REGION Network 6: Programmnummer gültig an den Schäumroboter
   //----
         L     #AB_KUKA_PGNO;
         T     #Prog_Nummer;
   //----
   // Partitätsbit auswerten
   //----
         X     #Temp_IO_Status.Output_To_Robot.A_SPS_PGNO.%X0;
         X     #Temp_IO_Status.Output_To_Robot.A_SPS_PGNO.%X1;
         X     #Temp_IO_Status.Output_To_Robot.A_SPS_PGNO.%X2;
         X     #Temp_IO_Status.Output_To_Robot.A_SPS_PGNO.%X3;
         X     #Temp_IO_Status.Output_To_Robot.A_SPS_PGNO.%X4;
         X     #Temp_IO_Status.Output_To_Robot.A_SPS_PGNO.%X5;
         X     #Temp_IO_Status.Output_To_Robot.A_SPS_PGNO.%X6;
         X     #Temp_IO_Status.Output_To_Robot.A_SPS_PGNO.%X7;
         =     #Temp_IO_Status.Output_To_Robot.A_SPS_PARITY;
   //----
   // Programmnummer an KUKA ablöschen, sobald sie erkannt wurde
   //----
         O(;
         A     #Temp_IO_Status.Input_From_Robot.E_KRC_PGNO_REQ;
         FN    #Temp_IO_Status.FHM_PRG_laeuft;
         );
         ON    #Temp_IO_Status.Input_From_Robot.E_KRC_PRO_ACT;
         ON    #Temp_IO_Status.Input_From_Robot.E_KRC_AUT_EXTERN;
         ON    #Temp_IO_Status.Anforderung_Automatik;
         O     #Temp_IO_Status.Input_From_Robot.E_KRC_MH_OPEN;
         JCN   strt;
         L     0;
         T     #Temp_IO_Status.A_SPS_PGNO;
         CLR;
         =     #Temp_IO_Status.Output_To_Robot.A_SPS_PARITY;
   //----
   strt: O(;
         L     #Temp_IO_Status.A_SPS_PGNO;
         L     0;
         >I;
         );
         =     #Temp_IO_Status.PrgNr_ok;

         A(;
         O     #IO_Button_MainPos;
         O     #IO_Button_Cleaning;
         O     #IN_Start_cycle;
         );
         A     #Temp_IO_Status.PrgNr_ok;
         L     S5T#100MS;
         SD    #IN_Timer_PGNO_Valid;
         A     #IN_Timer_PGNO_Valid;
         S     #Temp_IO_Status.Output_To_Robot.A_SPS_PGNO_VALID;

         A     #Temp_IO_Status.Output_To_Robot.A_SPS_PGNO_VALID;
         L     S5T#300MS;
         SE    #IN_Timer_Imp_ExtStart;

         A     #IN_Timer_Imp_ExtStart;
         =     #Temp_IO_Status.HM_Ext_Start;

   //    O     #Temp_IO_Status.HM_Ext_Start
   //    O     #Temp_IO_Status.Output_To_Robot.A_SPS_EXT_START
   //    =     #Temp_IO_Status.Output_To_Robot.A_SPS_EXT_START

         O(;
         A     #Temp_IO_Status.Output_To_Robot.A_SPS_EXT_START;
         FN    #Temp_IO_Status.FHM_PrgNr_gueltig;
         );
         O     #Temp_IO_Status.Input_From_Robot.E_KRC_APPL_RUN;
         ON    #Temp_IO_Status.Input_From_Robot.E_KRC_PRO_ACT;
         ON    #Temp_IO_Status.Input_From_Robot.E_KRC_AUT_EXTERN;
         R     #Temp_IO_Status.Output_To_Robot.A_SPS_PGNO_VALID;
   //-------------------------
         L     #Temp_IO_Status.A_SPS_PGNO;
         T     #Temp_IO_Status.Output_To_Robot.A_SPS_PGNO;
END_REGION

REGION Network 7: Signals MH
         A     #IN_Release_move_MC;
         =     #Temp_IO_Status.Output_To_Robot.A_SPS_DIRELMOVEMC;

         A     #IN_Shotrelease;
         =     #Temp_IO_Status.Output_To_Robot.A_SPS_READY_FOR_SHOT;

         A     #IN_Shotend;
         =     #Temp_IO_Status.Output_To_Robot.A_SPS_SHOTEND;

         A     #IN_OM_service;
         =     #Temp_IO_Status.Output_To_Robot.A_SPS_SERVICE;
END_REGION

REGION Network 8: Programmabbruch (Automatisches HP fahren)
         ON    #IN_Auto_Stop_quitt;
         O(;
         A     #IN_FLT_Group_1;
         A     #IN_Cycle_running;
         );
         A     #Temp_IO_Status.Input_From_Robot.E_KRC_AUT_EXTERN;
         AN    #Temp_IO_Status.Input_From_Robot.E_KRC_IN_HOME;
         AN    #Temp_IO_Status.Input_From_Robot.E_KRC_IN_MAINPOS;
         S     #Temp_IO_Status.Output_To_Robot.A_SPS_INTERRUPT;

         A     #Temp_IO_Status.Input_From_Robot.E_KRC_IN_HOME;
         R     #Temp_IO_Status.Output_To_Robot.A_SPS_INTERRUPT;
END_REGION

REGION Network 9: Ausgänge zum Roboter schreiben
         NOP   0;
   //
         L;
         LAR2;
         L     #IN_PW_INOUT;
         SLD   3;
         LAR1;
   //
         L     3;  // Länge der Ausgangsworte
   Palp: T     #Schleifenzaehler;
   //
         L     LW [ AR2 , P#30.0 ];  // Wert im Datenbaustein
         T     PQW [AR1,P#0.0];  // Ausgangswort
   //
         +AR1  P#2.0;
         +AR2  P#2.0;
   //
         L     #Schleifenzaehler;
         LOOP  Palp;
END_REGION

REGION Network 10: Daten sichern
   //----
         CALL  BLKMOV
         ( SRCBLK  := #Temp_IO_Status,
           RET_VAL := #ERROR_CODE,
           DSTBLK  := #Anyzeiger
         );
   //----
END_REGION
END_FUNCTION

FUNCTION "FC1910_IF_ABB" : Void   // FC1910, STL
TITLE = Interface foaming robot
{ S7_Optimized_Access := 'FALSE' }
AUTHOR : KT242
FAMILY : RS_KK
NAME : SS_ABB
VERSION : 2.1
   VAR_INPUT
      IN_PW_Ein_Ausgaenge : Int;   // Erste Adresse der Eingänge/ Ausgänge an/ vom Roboter
      IN_Reset_fault_Fkt : Bool;   // Signal zum quittieren der Störungen innerhalb der einzelnen Funktionsbausteine
      IN_Steuerspannung : Bool;   // Signal für eine Verzögerung der Ansteuerung der Umrichter (Schutz nach Not-Aus)
      IN_Zyklus_Laeuft : Bool;   // Signal das der Zyklus der Schäummaschine läuft
      IN_Zyklus_KLZ1_Laeuft : Bool;   // Signal das die Kreislaufzeit 1 der Schäummaschine läuft
      IN_Zyklus_KLZ3_Laeuft : Bool;   // Signal das die Kreislaufzeit 3 der Schäummaschine läuft
      IN_Zyklus_Schuss_laeuft : Bool;   // Signal das der Schuss läuft
      IN_Imp_Schussende : Bool;   // Signal das ein Teilschuss beendet wurde
      IN_Imp_Prog_Letzter_TS : Bool;   // Signal für das Ende des letzten Teilschusses eines Schäumprogrammes
      IN_Betriebsart_Automatik : Bool;   // Foaming machine in automatic mode
      IN_MK_Automatik : Bool;   // Eingang Mischkopf- Bedienpult befindet sich in der Stellung "Auto"
      IN_Anf_Flucht : Bool;   // Anforderung an den Roboter für eine Fluchtbewegung
      IN_Auto_Stop_quittiert : Bool;   // Automatikbetrieb kann gestartet werten, Automatik- Stopp ist quittiert
      IN_Zyklus_Freigabe : Bool;   // Die Freigabe zum Starten des Schäumzyklusses aus dem Zyklusbaustein steht an
      IN_Zyklus_Max_Wartezeit : Bool;   // Es wurde dir maximale Wartezeit nach KLZ 1 oder 3 überschritten
      IN_Start_Prog_Imp : Bool;   // Impulssignal zum Starten des Datenaustausches zum Roboter
      IN_FRG_Datatransfer : Bool;   // Freigabe zur Datenübertragung an den Roboter und zum anfahren der Vorposition
      IN_FRG_von_PU : Bool;   // Freigabe zum verfahren der Schäumbahn innerhalb des Formträgers
      IN_Anwahl_Mit_Shotware : Bool;   // Anwahl wenn der Roboter mit der Option Shotware betrieben wird
      IN_Anwahl_Mit_Tracking : Bool;   // Anwahl wenn der Roboter mit der Option Conveyer-Tracking betrieben wird
      IN_Timer_Auto_ein_Track : Timer;   // Timer für das Überprüfen des Trackingsignale doRobWaitWobj
      IN_Timer_Auto_ein : Timer;   // Timer für das automatische einschalten des Roboters
      IN_Timer_Verz_Handanwahl : Timer;   // Timer für das Verzögern des Motoren Ausschaltens bei Handanwahl
      IN_Timer_Auto_aus : Timer;   // Timer für das automatische ausschalten des Roboters
      IN_Timer_Fluchtprog : Timer;   // Timer für die Verlängereung des Signals für die Anforderung der Föuchtbewegung
      IN_Timer_Start_Verz : Timer;   // Timer zur Verzögerung des Programstartes nach Motoren ein
      IN_Timer_Start_Main_Verz : Timer;   // Timer zur Verzögerung des Programstartes Fahrt von Wartungspos->HP
      IN_Schusszeit : Word;   // Für den nächsten Eintrag benötigte Schußzeit
   END_VAR
   VAR_IN_OUT
      IO_Status : "ABB_IRC6_State";   // Speichern der Roboter- Zustände für das Programm
      IO_Fault : "General_Faults";
      IO_NewFault : Bool;
      IO_FaultLevel_1 : Bool;
      IO_FaultLevel_2 : Bool;
      IO_FaultLevel_3 : Bool;
   END_VAR
   VAR_TEMP
      Temp_IO_Status : "ABB_IRC6_State";   // Temporärer Roboter- Status für die interne Bearbeitung des Bausteins
      Temp_IO_Fault : "General_Faults";
      ERROR_CODE : Int;   // Error state of systemfunction "BLKMOV" Blockmove
      Anypointer1 : ANY;   // Pointer to copy thr array "IO_Status" and "Temp_IO_Status"
      Anypointer2 : ANY;   // Pointer to copy thr array "IO_Status" and "Temp_IO_Status"
      Adresse_im_Baustein : DWord;   // and the start adress within the program block
      Schleifenzaehler : Int;   // Zwischenmerker für die Schleifenzähler der verschiedenen Anwendungen
      Formen : Byte;   // Zwischenmerker für die Anzahl der aktuellen Formen
      Zeiten : Byte;   // Zwischenmerker für die Anzahl der aktuellen Zeiten
      Start_noetig : Bool;   // Zwischenmerker das das Starten des Roboters von Grund auf angefordert wird
      Imp_Roboter_in_Homepos : Bool;   // Impulsmerker das sich der Roboter in die Homeposition bewegt hat
      HM_Roboter_im_Programm : Bool;   // hilfsmerker für die Erkennung der Startsequenz
      Imp_Prog_n_Teilschuss : Bool;   // Impulsmerker für das Übertragen des nächsten Verfahrprogrammes
      Merker_Stoerung_Rob : Byte;   // Zwischenmerker für die Darstellung der Störungen
      Merker_StNrRob_OUT : Word;   // Zwischenmerker für die Darstellung der Störungen
      Merker_TimeNr : Byte;   // Zwischenmerker für den aktuellen TS in der aktuellen Form
      TestPAW : Word;
      RefMerk : DWord;
   END_VAR
BEGIN

REGION Network 1: Saved data integration
         LAR1;
         L;
         LAR2;
   //
         L     16#1002;  // Bytes
         T     W[AR1, P#0.0];
         L     60;  // Amount of bytes
         T     W[AR1, P#2.0];
         L     W [ AR2 , P#0.0 ];  // Block no,
         T     W[AR1, P#4.0];
         L     D [ AR2 , P#2.0 ];  // Startadress of datas
         T     D[AR1, P#6.0];
   //
         CALL  BLKMOV
         ( SRCBLK  := #Anypointer1,
           RET_VAL := #ERROR_CODE,
           DSTBLK  := #Temp_IO_Status
         );
   //
   //
         LAR1;
         L;
         LAR2;
   //
         L     16#1002;  // Bytes
         T     W[AR1, P#0.0];
         L     4;  // Amount of bytes
         T     W[AR1, P#2.0];
         L     W [ AR2 , P#0.0 ];  // Block no,
         T     W[AR1, P#4.0];
         L     D [ AR2 , P#2.0 ];  // Startadress of datas
         T     D[AR1, P#6.0];
   //
         CALL  BLKMOV
         ( SRCBLK  := #Anypointer2,
           RET_VAL := #ERROR_CODE,
           DSTBLK  := #Temp_IO_Fault
         );
   //
END_REGION

REGION Network 2: Ausgänge von dem Roboter in die Steuerung laden
         L;
         LAR2;
         L     #IN_PW_Ein_Ausgaenge;
         SLD   3;
         LAR1;
   //
         L     8;  // Anzahl der Eingangsworte
   Pelp: T     #Schleifenzaehler;
   //
         L     PIW[AR1, P#0.0];  // Eingangsswort
         T     LW[AR2, P#34.0];  // Ausgänge im UDT
   //
         +AR1  P#2.0;
         +AR2  P#2.0;
   //
         L     #Schleifenzaehler;
         LOOP  Pelp;
END_REGION

REGION Network 3: Störung
         A     #IN_Reset_fault_Fkt;
         R     #Temp_IO_Status.STG_System;
         R     #Temp_IO_Status.Fault_from_system;
         R     #Temp_IO_Fault.FLT_System;
         R     #Temp_IO_Fault.FLT_Wrong_Shot_time;
         R     #Temp_IO_Fault.FLT_Wrong_Prog_No;
         R     #Temp_IO_Fault.FLT_Wrong_MC_No;
         R     #Temp_IO_Fault.FLT_Prog_stopped;
         R     #Temp_IO_Fault.FLT_Fuse;
   //
         A     #IN_Reset_fault_Fkt;
         A     #Temp_IO_Status.Output.doSysError;
         =     #Temp_IO_Status.Input.diResetError;
   //
         A     #IN_Reset_fault_Fkt;
         A     #Temp_IO_Status.Output.doEmStop_Akt;
         =     #Temp_IO_Status.Input.diResetEstop;
   //
         A     #Temp_IO_Status.Auto_mode_requested;
         A     #IN_Timer_Auto_ein;
         A     #Temp_IO_Status.Output.doSysError;
         S     #Temp_IO_Status.STG_System;
   //
         AN    #Temp_IO_Status.STG_System;
         AN    #Temp_IO_Status.Fault_from_system;
         R     #Temp_IO_Status.Fault_observed;
   //
         O     #Temp_IO_Status.STG_System;
         O     #Temp_IO_Status.Fault_from_system;
         A     #Temp_IO_Status.Output.doIRBinAuto;
         S     #Temp_IO_Status.Fault_observed;
   //
         AN    #Temp_IO_Status.Fault_observed;
         =     #Temp_IO_Status.Interface_OK;
END_REGION

REGION Network 4: Anwahl Automatik/Hand anfordern
         A     #IN_Steuerspannung;
         A(;
         O     #IN_MK_Automatik;
         O     #Temp_IO_Status.Input.diMaintToHomeP;
   //      O     #Temp_IO_Status.Input.diServiceShot
         );
         A     #IN_Auto_Stop_quittiert;
         A     #Temp_IO_Status.Output.doIRBinAuto;
         A     #Temp_IO_Status.Interface_OK;
         AN(;
         A     #IN_Anwahl_Mit_Tracking;
         A     #Temp_IO_Status.Output.doIRBSyncWobj;
         AN    #IN_Zyklus_Freigabe;
         A     #IN_Timer_Auto_ein_Track;
         );
         A     #IN_Betriebsart_Automatik;
         AN    #Temp_IO_Status.Output.doSafeZoneActiv;
         =     #Temp_IO_Status.Auto_mode_requested;
   //
         AN    #Temp_IO_Status.Auto_mode_requested;
         L     S5T#2S;
         SP    #IN_Timer_Auto_aus;
   //
         A     #IN_Timer_Auto_aus;
         O(;
         A     #Temp_IO_Status.Output.doSafeZoneActiv;
         A     #Temp_IO_Status.Output.doIRBinAuto;
         );
         =     #Temp_IO_Status.Manual_mode_requested;
END_REGION

REGION Network 5: Entscheidung über die Art des Starts
         ON    #Temp_IO_Status.Output.doIRBinAuto;
         O     #Temp_IO_Status.Output.doSysError;
         S     #Temp_IO_Status.Robot_not_in_Auto;
   //
         O     #Temp_IO_Status.Output.doIRBInHome;
         FP    #Temp_IO_Status.HF_Robot_not_in_Auto;
         =     #Imp_Roboter_in_Homepos;
         O     #Temp_IO_Status.Input.diStartCycle;
         O     #Temp_IO_Status.Input.diMaintToHomeP;
         O     #Imp_Roboter_in_Homepos;
         A     #Temp_IO_Status.Output.doIRBinAuto;
         R     #Temp_IO_Status.Robot_not_in_Auto;
   //
         A     #Temp_IO_Status.Output.doIRBInMaintP;
         O(;
         A     #Temp_IO_Status.Input.diBreak;
         AN    #Temp_IO_Status.Output.doIRBOutRangMC;
         );
         O(;
         A     #Temp_IO_Status.Input.diJumpConveyer;
         A     #Temp_IO_Status.Output.doIRBOutRangMC;
         );
         =     #HM_Roboter_im_Programm;
   //
         A     #HM_Roboter_im_Programm;
         AN    #Temp_IO_Status.Robot_not_in_Auto;
         AN(;
         A     #IN_Anwahl_Mit_Tracking;
         A     #Temp_IO_Status.Output.doIRBSyncWobj;
         );
         A     #Temp_IO_Status.Auto_mode_requested;
         =     #Temp_IO_Status.Robot_processing_prog;
END_REGION

REGION Network 6: Anwahl Automatik
         A     #Temp_IO_Status.Auto_mode_requested;
         AN    #Temp_IO_Status.Output.doMotorOn;
         A     #Temp_IO_Status.Output.doMotorOff;
         AN    #Temp_IO_Status.Output.doCycleOn;
         R     #Temp_IO_Status.Input.diMotorOff;
         L     S5T#2S;  // S5T#1S
         SD    #IN_Timer_Start_Verz;
         A     #IN_Timer_Start_Verz;
         S     #Temp_IO_Status.Input.diMotorOn;
   //
         A     #Temp_IO_Status.Auto_mode_requested;
         A     #Temp_IO_Status.Output.doMotorOn;
         AN    #Temp_IO_Status.Output.doMotorOff;
         AN    #Temp_IO_Status.Output.doCycleOn;
         R     #Temp_IO_Status.Input.diMotorOn;
         =     #Start_noetig;
   //

         A     #Start_noetig;
         A     #Temp_IO_Status.Robot_processing_prog;
         S     #Temp_IO_Status.Input.diStartProg;
         A     #Start_noetig;
         AN    #Temp_IO_Status.Robot_processing_prog;
         L     s5t#500ms;
         SD    #IN_Timer_Start_Main_Verz;  //Problem wenn Roboter fährt von Maint. Pos->Homepos bleiben Motoren ein abe Programm stoppt
         A     #IN_Timer_Start_Main_Verz;
         S     #Temp_IO_Status.Input.diStartMain;

   //
         A     #Temp_IO_Status.Auto_mode_requested;
         A     #Temp_IO_Status.Output.doMotorOn;
         AN    #Temp_IO_Status.Output.doMotorOff;
         A     #Temp_IO_Status.Output.doCycleOn;
         R     #Temp_IO_Status.Input.diStartProg;
         R     #Temp_IO_Status.Input.diStartMain;
         =     #Temp_IO_Status.Auto_accepted;
   //
         A     #Temp_IO_Status.Auto_accepted;
         L     S5T#500MS;
         SD    #IN_Timer_Auto_ein;
         L     S5T#2S;
         SD    #IN_Timer_Auto_ein_Track;
   //
         ON    #Temp_IO_Status.Auto_mode_requested;
         O     #Temp_IO_Status.Output.doSysError;
         R     #Temp_IO_Status.Input.diMotorOn;
         R     #Temp_IO_Status.Input.diStartProg;
         R     #Temp_IO_Status.Input.diStartMain;
END_REGION

REGION Network 7: Anwahl Hand
         A     #Temp_IO_Status.Output.doMotorOn;
         AN    #Temp_IO_Status.Output.doMotorOff;
         O     #Temp_IO_Status.Output.doCycleOn;
         A     #Temp_IO_Status.Manual_mode_requested;
         S     #Temp_IO_Status.Input.diStopProg;
         L     S5T#1S;
         SD    #IN_Timer_Verz_Handanwahl;
   //
         A     #IN_Timer_Verz_Handanwahl;
         A     #Temp_IO_Status.Manual_mode_requested;
         A     #Temp_IO_Status.Output.doMotorOn;
         AN    #Temp_IO_Status.Output.doMotorOff;
         AN    #Temp_IO_Status.Output.doCycleOn;
         R     #Temp_IO_Status.Input.diStopProg;
         S     #Temp_IO_Status.Input.diMotorOff;
   //
         A     #Temp_IO_Status.Manual_mode_requested;
         AN    #Temp_IO_Status.Output.doMotorOn;
         A     #Temp_IO_Status.Output.doMotorOff;
         AN    #Temp_IO_Status.Output.doCycleOn;
         R     #Temp_IO_Status.Input.diMotorOff;
   //
         ON    #Temp_IO_Status.Manual_mode_requested;
         O     #Temp_IO_Status.Output.doSysError;
         R     #Temp_IO_Status.Input.diStopProg;
         R     #Temp_IO_Status.Input.diMotorOff;
END_REGION

REGION Network 8: Fluchtprogramm starten
         A     #IN_Anf_Flucht;
         AN    #Temp_IO_Status.Output.doStopFormPLC;
         S     #Temp_IO_Status.Escape_program;
         S     #Temp_IO_Status.Input.diInterrupt;
         L     S5T#3S;
         SE    #IN_Timer_Fluchtprog;
   //
         ON    #IN_Timer_Fluchtprog;
         R     #Temp_IO_Status.Escape_program;
         R     #Temp_IO_Status.Input.diInterrupt;
END_REGION

REGION Network 9: Freigabe Schäumzyklus / Reset / Ende
         A     #IN_Zyklus_Freigabe;
         AN    #IN_Anf_Flucht;
         A     #Temp_IO_Status.Auto_accepted;
         =     #Temp_IO_Status.Freigabe_Schaeumzyklus;
   //
         A     #Temp_IO_Status.Freigabe_Schaeumzyklus;
         AN    #IN_Zyklus_Max_Wartezeit;
         JC    spgl;
         JU    res;
END_REGION

REGION Network 10: Sprungleiste Datenübertragung
   spgl: L     #Temp_IO_Status.Stepnumber;
   //
         JL    del;
         JU    strt;  //  0: Warten auf Start
         JU    wrtt;  //  1: Warten auf Schusszeiten
         JU    aMld;  //  2: Anzahl Teilformen
         JU    zygo;  //  3: Roboterzyklus Datenaustausch starten
         JU    aPr;  //  4: Aktuelles Verfahrprogramm bestimmen
         JU    dglt;  //  5: Daten gültig setzen
         JU    dan0;  //  6: Daten gültig rücksetzen
         JU    Nmld;  //  7: Noch eine Form schäumen??
         JU    vpos;  //  8: Vorposition abwarten
         JU    ssig;  //  9: Schäumsignale ausgeben
   del:  JU    res;
   //
   res:  L     0;
         T     #Temp_IO_Status.Mould_Number;
         T     #Temp_IO_Status.Offset_of_Shottime;
         T     #Temp_IO_Status.Stepnumber;
         T     #Temp_IO_Status.Input.GIMCNo;
         T     #Temp_IO_Status.Input.GIProgNo1;
         T     #Temp_IO_Status.Input.GIShotTX1;
         L     1;
         T     #Temp_IO_Status.Time_Nummer;
   //
         SET;
         R     #Temp_IO_Status.Input.diStartCycle;
         R     #Temp_IO_Status.Input.diReadProgNo;
   //      R     #Temp_IO_Status.Input.diShotDigIn
   //
         R     #Temp_IO_Status.Input.giMouldCodeBit0;
         R     #Temp_IO_Status.Input.giMouldCodeBit1;
   //
         R     #Temp_IO_Status.Release_foaming;
         R     #Temp_IO_Status.Shot_time_received;
         R     #Temp_IO_Status.Data_transmitted;
         R     #Temp_IO_Status.Motion_prog01_existing;
         R     #Temp_IO_Status.Motion_prog02_existing;
         R     #Temp_IO_Status.Motion_prog03_existing;
         R     #Temp_IO_Status.HFShotDigOut_open_MH;
         R     #Temp_IO_Status.doShotDigOut_open_MH;
         JU    WRSZ;
END_REGION

REGION Network 11: Schritt 0: Start Schäumzyklus
   strt: ON    #IN_Start_Prog_Imp;
         JC    WRSZ;
   //
   //      L     0                    // Beginnend bei Wort Null
   //      LAR1                       // Adresse für Schußzeit im DB
   //
   //      L     60                   // Anzahl der Schußzeiten
   //clrF: NOP 0                      // Öffnen des Schußzeitenbausteins
   //      T     #Schleifenzaehler
   //
   //      AUF   #IN_Schusszeit
   //      L     0
   //      T DBW [ AR1 , P#0.0 ]
   //
   //      +AR1  P#2.0
   //
   //      L     #Schleifenzaehler    // Wenn Schleifenzähler <> 0
   //      LOOP  clrF                 // Schleife erneut durchlaufen
   //
   // Ablöschen der Verfahrprogramme:
   //
   //      L     320                  // Beginnend bei Datenwot 320
   //      SLD   3
   //      LAR1                       // Adresse für Verfahrprogramme im DB
   //
   //      L     8                    // Anzahl der Verfahrprogramme
   //clrV: NOP 0                      // Öffnen des Schußzeitenbausteins
   //      T     #Schleifenzaehler
   //
   //      AUF   #IN_Schusszeit
   //      L     0
   //      T DBW [ AR1 , P#0.0 ]
   //
   //      +AR1  P#2.0
   //
   //      L     #Schleifenzaehler    // Wenn Schleifenzähler <> 0
   //      LOOP  clrV                 // Schleife erneut durchlaufen
   //
         L     #Temp_IO_Status.Stepnumber;
         +     1;
         T     #Temp_IO_Status.Stepnumber;
         JU    WRSZ;
END_REGION

REGION Network 12: Schritt 1: Warten auf Schusszeiten
   wrtt: NOP   0;
         L     #IN_Schusszeit;
         L     0;
         <>D;
         ON    #IN_Anwahl_Mit_Shotware;
         A(;
         O(;
         L     #Temp_IO_Status.Robot_ProgNo_Mould_1;
         L     0;
         <>D;
         );
         O(;
         L     #Temp_IO_Status.Robot_ProgNo_Mould_2;
         L     0;
         <>D;
         );
         O(;
         L     #Temp_IO_Status.Robot_ProgNo_Mould_3;
         L     0;
         <>D;
         );
         );
         JCN   WRSZ;
   //
         L     #Temp_IO_Status.Stepnumber;
         +     1;
         T     #Temp_IO_Status.Stepnumber;
         JU    WRSZ;
END_REGION

REGION Network 13: Schritt 2: Anzahl Verfahrwege festlegen
   aMld: NOP   0;
   //_________________________________________________
   // Verfahrweg für die Form Nr.3 ist vorhanden
         A(;
         L     #Temp_IO_Status.Robot_ProgNo_Mould_3;
         L     0;
         ==D;
         );
         JC    F2;
   //
         SET;
         S     #Temp_IO_Status.Motion_prog01_existing;
         S     #Temp_IO_Status.Motion_prog02_existing;
         S     #Temp_IO_Status.Motion_prog03_existing;
         S     #Temp_IO_Status.Input.giMouldCodeBit0;
         S     #Temp_IO_Status.Input.giMouldCodeBit1;
         JU    MCNr;
   //_________________________________________________
   // Verfahrweg für die Form Nr.2 ist vorhanden
   F2:   O(;
         L     #Temp_IO_Status.Robot_ProgNo_Mould_2;
         L     0;
         ==D;
         );
         JC    F3;
   //
         SET;
         S     #Temp_IO_Status.Motion_prog01_existing;
         S     #Temp_IO_Status.Motion_prog02_existing;
         S     #Temp_IO_Status.Input.giMouldCodeBit1;
         JU    MCNr;
   //_________________________________________________
   // Verfahrweg für die Form Nr.1 ist vorhanden
   F3:   O(;
         L     #Temp_IO_Status.Robot_ProgNo_Mould_1;
         L     0;
         ==D;
         );
         JC    MCNr;
   //
         SET;
         S     #Temp_IO_Status.Motion_prog01_existing;
         S     #Temp_IO_Status.Input.giMouldCodeBit0;
   //_______________________________________________
   //
   MCNr: NOP   0;
         L     #Temp_IO_Status.MC_Place_Number;
         T     #Temp_IO_Status.Input.GIMCNo;
   //
         L     #Temp_IO_Status.Stepnumber;
         +     1;
         T     #Temp_IO_Status.Stepnumber;
         JU    WRSZ;
END_REGION

REGION Network 14: Schritt 3: Zyklusstart für Datenaustausch setzen
   zygo: NOP   0;
   //
         A     #IN_FRG_Datatransfer;
         S     #Temp_IO_Status.Input.diStartCycle;
         JCN   WRSZ;
   //
         L     #Temp_IO_Status.Stepnumber;
         +     1;
         T     #Temp_IO_Status.Stepnumber;
         JU    WRSZ;
END_REGION

REGION Network 15: Schritt 4: Aktuelle Formnummer festlegen
   aPr:  NOP   0;
   //
         A     #Temp_IO_Status.Motion_prog01_existing;
         JCN   a2FT;
         SET;
         R     #Temp_IO_Status.Motion_prog01_existing;
   //
         L     #Temp_IO_Status.Robot_ProgNo_Mould_1;
         CAW;
         T     #Temp_IO_Status.Input.GIProgNo1;
   //
         JU    aPre;
   ///
   a2FT: A     #Temp_IO_Status.Motion_prog02_existing;
         JCN   a3FT;
         SET;
         R     #Temp_IO_Status.Motion_prog02_existing;
   //
         L     #Temp_IO_Status.Robot_ProgNo_Mould_2;
         CAW;
         T     #Temp_IO_Status.Input.GIProgNo1;
   //
         JU    aPre;
   //
   a3FT: A     #Temp_IO_Status.Motion_prog03_existing;
         JCN   aPre;
         SET;
         R     #Temp_IO_Status.Motion_prog03_existing;
   //
         L     #Temp_IO_Status.Robot_ProgNo_Mould_3;
         CAW;
         T     #Temp_IO_Status.Input.GIProgNo1;
   //
         JU    aPre;
   //
   aPre: L     #Temp_IO_Status.Stepnumber;
         +     1;
         T     #Temp_IO_Status.Stepnumber;
         JU    WRSZ;
END_REGION

REGION Network 16: Schritt 5: Daten gültig setzen
   dglt: S     #Temp_IO_Status.Input.diReadProgNo;
   //
         L     #Temp_IO_Status.Stepnumber;
         +     1;
         T     #Temp_IO_Status.Stepnumber;
         JU    WRSZ;
END_REGION

REGION Network 17: Schritt 6: Wenn Datenanforderung rückgesetzt-Daten gültig löschen
   dan0: AN    #Temp_IO_Status.Output.doProgNoReaded;
         JC    WRSZ;
         R     #Temp_IO_Status.Input.diReadProgNo;
   //
         L     #Temp_IO_Status.Stepnumber;
         +     1;
         T     #Temp_IO_Status.Stepnumber;
         JU    WRSZ;
END_REGION

REGION Network 18: Schritt 7: Warten bis Roboter bereit zum Empfang für neue Daten
   Nmld: NOP   0;
   //
         A     #Temp_IO_Status.Output.doProgNoReaded;
         JC    WRSZ;
   //
         AN    #Temp_IO_Status.Motion_prog01_existing;
         AN    #Temp_IO_Status.Motion_prog02_existing;
         AN    #Temp_IO_Status.Motion_prog03_existing;
         JC    shot;
   //
         L     4;  // 4: Nächstes Verfahrprogramm
         T     #Temp_IO_Status.Stepnumber;
         JU    WRSZ;
   //
   shot: L     #Temp_IO_Status.Stepnumber;
         +     1;
         T     #Temp_IO_Status.Stepnumber;
         JU    WRSZ;
END_REGION

REGION Network 19: Schritt 8: Warten bis Homeposition verlassen wurde
   vpos: NOP   0;
         A     #Temp_IO_Status.Output.doIRBInHome;
         JC    WRSZ;
   //
         R     #Temp_IO_Status.Input.diStartCycle;

         L     #Temp_IO_Status.Stepnumber;
         +     1;
         T     #Temp_IO_Status.Stepnumber;
         JU    WRSZ;
END_REGION

REGION Network 20: Schritt 9: Warten bis Zyklusende gemeldet wird
   // An dieser Stelle wird nur direkt der Schäumvorgang abgewickelt. 
   // Anlagenspezifische Signale wie z.B. der MK-Reiniger sollten besser extern 
   // belegt werden. Ideal ist die Belegung vor dem Aufruf der Funktion FC 113, da 
   // dann die Daten im gleichen SPS-Zyklus an die Peripherie übertragen werden.
   ssig: NOP   0;
         A     #IN_FRG_von_PU;  // Shot release from foaming cycle
         A(;
         O     #Temp_IO_Status.Input.diShotDigIn;
         ON    #Temp_IO_Status.Output.doShotDigOut;
         );
         =     #Temp_IO_Status.Input.diShotDigIn;
   //
   // Aus Sicherheitsgründen: Flankenabfrage des MK - öffnens
   //
         A     #Temp_IO_Status.Output.doShotDigOut;
         FP    #Temp_IO_Status.HFShotDigOut_open_MH;
         S     #Temp_IO_Status.doShotDigOut_open_MH;
   //
         O     #IN_Imp_Schussende;
         ON    #IN_Zyklus_Laeuft;
         R     #Temp_IO_Status.doShotDigOut_open_MH;

   // Zyklusende mit Homeposition
         AN    #Temp_IO_Status.Output.doCycleEnd;
         JC    WRSZ;
   //
         L     #Temp_IO_Status.Stepnumber;
         +     1;
         T     #Temp_IO_Status.Stepnumber;
         JU    WRSZ;
END_REGION

REGION Network 21: Aktuelle Schusszeit an den Roboter schreiben
   // An dieser Stelle wir dem Roboter immer die für den nächsten Teilschuss aktuelle 
   // Schusszeit zur verfügung gestellt!
   WRSZ: NOP   0;
   //
   // Reset TeileschussNr wenn eine neue Form begonnen wird
   //
         A     #IN_Imp_Prog_Letzter_TS;
         JCN   SZRS;
         L     1;
         T     #Temp_IO_Status.Time_Nummer;
   SZRS: NOP   0;
   //
         A     #IN_Zyklus_Schuss_laeuft;
         A     #IN_Zyklus_Laeuft;
         FP    #Temp_IO_Status.HF_next_partshot;
         =     #Imp_Prog_n_Teilschuss;
   //
         A     #Imp_Prog_n_Teilschuss;
         JCN   SZ01;
   //
   // Bestimmen des nächsten Teilschusses
   //
         L     #Temp_IO_Status.Time_Nummer;
         L     1;
         +I;
         T     #Temp_IO_Status.Time_Nummer;
   //
   SZ01: NOP   0;
   //
   // Bestimmen der aktuellen Form für die Zeiten
   //
         L     0;
         AN    #Temp_IO_Status.Output.goMouldActBit0;
         A     #Temp_IO_Status.Output.goMouldActBit1;
         JCN   SZ02;
         L     40;
   SZ02: NOP   0;
   //
         A     #Temp_IO_Status.Output.goMouldActBit0;
         A     #Temp_IO_Status.Output.goMouldActBit1;
         JCN   SZ03;
         L     80;
   SZ03: NOP   0;
         T     #Temp_IO_Status.Offset_of_Shottime;
   //
         L     0;
         L     #Temp_IO_Status.Time_Nummer;
         ==I;
         JC    SZ04;
         L     1;
         -I;
   SZ04: NOP   0;
         T     #Merker_TimeNr;
   //
         L     #Merker_TimeNr;
         L     2;
         *I;
         L     #Temp_IO_Status.Offset_of_Shottime;
         +I;
         SLD   3;
         LAR1;
   //
   // aktuelle Schusszeit an Roboter transferieren
   //      AUF   #IN_Schusszeit
   //      L DBW [ AR1 , P#0.0 ]
   //      TAW

         L     #IN_Schusszeit;
         T     #Temp_IO_Status.Input.GIShotTX1;
END_REGION

REGION Network 22: PAW schreiben
         NOP   0;
   //
   //      L     400
   //      T     #TestPAW

         L;
         LAR2;
         L     #IN_PW_Ein_Ausgaenge;
         SLD   3;
         LAR1;
   //
         L     8;  // Länge der Ausgangsworte
   Palp: T     #Schleifenzaehler;
         L     LW[AR2, P#18.0];  // Wert im Datenbaustein
         T     PQW[AR1, P#0.0];  // Ausgangswort
   //
         +AR1  P#2.0;
         +AR2  P#2.0;
   //
         L     #Schleifenzaehler;
         LOOP  Palp;
END_REGION

REGION Network 23: Roboter Störungsnummer ausgeben
         L;
         LAR1;
   //
   // Aktuelle Meldungen ablöschen
   //
         L     5;  // Länge der Ausgangsworte
   ROBM: T     #Schleifenzaehler;
   //
         L     0;  // Wert im Datenbaustein
         T     LW[AR1, P#50.0];  // Ausgangswort
   //
         +AR1  P#2.0;
   //
         L     #Schleifenzaehler;
         LOOP  ROBM;
   //
         A(;
         L     0;
         L     #Temp_IO_Status.Output.GOError;
         <=D;
         );
         A(;
         L     17;
         <D;
         );
         JC    WA01;
   //
         A(;
         L     16;
         L     #Temp_IO_Status.Output.GOError;
         <D;
         );
         A(;
         L     33;
         <D;
         );
         JC    WA02;
   //
         A(;
         L     32;
         L     #Temp_IO_Status.Output.GOError;
         <D;
         );
         A(;
         L     49;
         <D;
         );
         JC    WA03;
   //
         A(;
         L     48;
         L     #Temp_IO_Status.Output.GOError;
         <D;
         );
         A(;
         L     65;
         <D;
         );
         JC    WA04;
   //
         A(;
         L     64;
         L     #Temp_IO_Status.Output.GOError;
         <D;
         );
         A(;
         L     81;
         <D;
         );
         JC    WA05;
   //_________________________________________________________________________
   //
   WA01: NOP   0;
         L     #Temp_IO_Status.Output.GOError;
         T     #Merker_Stoerung_Rob;
   //
         CALL  "FC107_Binär->Bit"
         ( IN_BinaerZahl := #Merker_Stoerung_Rob,
           OUT_BitZahl   := #Merker_StNrRob_OUT
         );
   //
         L;
         LAR1;
   //
         L     #Merker_StNrRob_OUT;  // Wert im Datenbaustein
         T     LW[AR1, P#50.0];  // Ausgangswort
         JU    WAEN;
   //
   WA02: NOP   0;
         L     #Temp_IO_Status.Output.GOError;
         L     16;
         -D;
         T     #Merker_Stoerung_Rob;
   //
         CALL  "FC107_Binär->Bit"
         ( IN_BinaerZahl := #Merker_Stoerung_Rob,
           OUT_BitZahl   := #Merker_StNrRob_OUT
         );
   //
         L;
         LAR2;
   //
         L     #Merker_StNrRob_OUT;  // Wert im Datenbaustein
         T     LW[AR2, P#52.0];  // Ausgangswort
         JU    WAEN;
   //
   WA03: NOP   0;
         L     #Temp_IO_Status.Output.GOError;
         L     32;
         -D;
         T     #Merker_Stoerung_Rob;
   //
         CALL  "FC107_Binär->Bit"
         ( IN_BinaerZahl := #Merker_Stoerung_Rob,
           OUT_BitZahl   := #Merker_StNrRob_OUT
         );
   //
         L;
         LAR2;
   //
         L     #Merker_StNrRob_OUT;  // Wert im Datenbaustein
         T     LW[AR2, P#54.0];  // Ausgangswort
         JU    WAEN;
   //
   WA04: NOP   0;
         L     #Temp_IO_Status.Output.GOError;
         L     48;
         -D;
         T     #Merker_Stoerung_Rob;
   //
         CALL  "FC107_Binär->Bit"
         ( IN_BinaerZahl := #Merker_Stoerung_Rob,
           OUT_BitZahl   := #Merker_StNrRob_OUT
         );
   //
         L;
         LAR1;
   //
         L     #Merker_StNrRob_OUT;  // Wert im Datenbaustein
         T     LW[AR1, P#56.0];  // Ausgangswort
         JU    WAEN;
   //
   WA05: NOP   0;
         L     #Temp_IO_Status.Output.GOError;
         L     64;
         -D;
         T     #Merker_Stoerung_Rob;
   //
         CALL  "FC107_Binär->Bit"
         ( IN_BinaerZahl := #Merker_Stoerung_Rob,
           OUT_BitZahl   := #Merker_StNrRob_OUT
         );
   //
         L;
         LAR1;
   //
         L     #Merker_StNrRob_OUT;  // Wert im Datenbaustein
         T     LW[AR1, P#58.0];  // Ausgangswort
   //
   WAEN: NOP   0;
END_REGION

REGION Network 24: Error handling
   //      O     XXXXXXXX
   //      S     #IO_FaultLevel_2

   //      O     xxxxxxxx
   //      S     #IO_FaultLevel_3

         O     #Temp_IO_Status.Output.doSysError;
         A     #Temp_IO_Status.Auto_mode_requested;
         AN    #Temp_IO_Fault.FLT_System;
         S     #Temp_IO_Fault.FLT_System;
         S     #IO_NewFault;

         O     #Temp_IO_Status.Meldungen.Rob_ST_17_32.FLT_No_019;
         A     #Temp_IO_Status.Auto_mode_requested;
         AN    #Temp_IO_Fault.FLT_Wrong_Prog_No;
         S     #Temp_IO_Fault.FLT_Wrong_Prog_No;
         S     #IO_NewFault;

         O     #Temp_IO_Status.Meldungen.Rob_ST_17_32.FLT_No_023;
         O     #Temp_IO_Status.Meldungen.Rob_ST_17_32.FLT_No_024;
         A     #Temp_IO_Status.Auto_mode_requested;
         AN    #Temp_IO_Fault.FLT_Wrong_Shot_time;
         S     #Temp_IO_Fault.FLT_Wrong_Shot_time;
         S     #IO_NewFault;

         O     #Temp_IO_Status.Meldungen.Rob_ST_17_32.FLT_No_022;
         O     #Temp_IO_Status.Meldungen.Rob_ST_33_48.FLT_No_044;
         A     #Temp_IO_Status.Auto_mode_requested;
         AN    #Temp_IO_Fault.FLT_Wrong_MC_No;
         S     #Temp_IO_Fault.FLT_Wrong_MC_No;
         S     #IO_NewFault;

         O     #Temp_IO_Status.Meldungen.Rob_ST_17_32.FLT_No_021;
         O     #Temp_IO_Status.Meldungen.Rob_ST_33_48.FLT_No_045;
         A     #Temp_IO_Status.Auto_mode_requested;
         AN    #Temp_IO_Fault.FLT_Prog_stopped;
         S     #Temp_IO_Fault.FLT_Prog_stopped;
         S     #IO_NewFault;

         O     #Temp_IO_Fault.FLT_System;
         O     #Temp_IO_Fault.FLT_Wrong_Shot_time;
         O     #Temp_IO_Fault.FLT_Wrong_Prog_No;
         O     #Temp_IO_Fault.FLT_Wrong_MC_No;
         O     #Temp_IO_Fault.FLT_Prog_stopped;
         S     #IO_FaultLevel_1;

         O     #Temp_IO_Fault.FLT_Fuse;
         S     #IO_FaultLevel_3;
END_REGION

REGION Network 25: Save data
         CALL  BLKMOV
         ( SRCBLK  := #Temp_IO_Status,
           RET_VAL := #ERROR_CODE,
           DSTBLK  := #Anypointer1
         );
   //
         CALL  BLKMOV
         ( SRCBLK  := #Temp_IO_Fault,
           RET_VAL := #ERROR_CODE,
           DSTBLK  := #Anypointer2
         );
   //
END_REGION
END_FUNCTION

FUNCTION "FC1920_IF_Fanuc" : Void   // FC1920, STL
TITLE = Interface to foaming robot
{ S7_Optimized_Access := 'FALSE' }
AUTHOR : KT242
NAME : IF_Fanuc
VERSION : 2.0
   VAR_INPUT
      IN_AdressRobIO : Hw_Io;   // Start Adress of Robot I/Os
      IN_ResetFaultFct : Bool;   // Signal to reset fault bits
      IN_ControlVoltage : Bool;   // Control voltage on
      IN_FoamingCycleRunning : Bool;   // Foaming cycle running
      IN_MHAutomatic : Bool;   // Key switch MH in automatic mode
      IN_RequestEscapeProg : Bool;   // Request escaping program
      IN_AutoStopOK : Bool;   // Automatic stop is ok
      IN_FuseSupplyOK : Bool;   // The fuse for power supply of robot is ok
      IN_EnableFoamingCycle : Bool;   // Enable signal for foaming cycle
      IN_ShotActive : Bool;   // Shot active
      IN_CycleMaxWaitingTime : Bool;   // Fault: maximum waiting time for shot
      IN_StartPulseDataExchang : Bool;   // Pulse start data transfer with robot
      IN_PulseShotEnd : Bool;   // Pulse part shot finished
      IN_EnableDataExchange : Bool;   // Enable data exchange with the robot
      IN_EnableShotFromPU : Bool;   // Enable shot from foaming machine
      IN_ConfigWithTracking : Bool;   // Configuration bit: robot with conveyor tracking
      IN_OtherRobotOnly : Bool;   // Only the other robot is activated for production
      IN_CleaningRequest : Bool;
      IN_PGNO_MainPos : Int;   // Programmnummer für Bewegung in Wartungsposition
      IN_PGNO_MainPos2 : Int;   // Programmnummer für Bewegung in Wartungsposition 2
      IN_PGNO_Cleaning : Int;   // Programmnummer für Bewegung zum Reinigen
      IN_PGNO_Testshot : Int;   // Programmnummer für Bewegung zur Testschussstation
      IN_TimerAutoOnTrack : Timer;   // Timer for monitoring the tracking signals doRobWaitWobj
      IN_TimerAutoOn : Timer;   // Timer for automatic switching on of the robot
      IN_TimerDelayManSelect : Timer;   // Delay timer for motor off when manual mode is selected
      IN_TimerAutoOFF : Timer;   // Timer for automatic switching off of the robot
      IN_TimerEscapeProg : Timer;   // Timer for requesting escape program
      IN_TimerStartDelay : Timer;   // Delay timer for program start after motor on
      IN_TimerFaultReset : Timer;   // Timer to set reset signal to robot
   END_VAR
   VAR_IN_OUT
      IO_Button_MainPos : Bool;   // Schalter Wartungsposition
      IO_Button_MainPos2 : Bool;   // Schalter Wartungsposition 2
      IO_Button_Cleaning : Bool;   // Schalter Reinigen
      IO_Button_Testshot : Bool;   // Schalter Testschuss
      IO_State_MainPos : Byte;   // Status Wartungsposition
      IO_State_MainPos2 : Byte;   // Status Wartungsposition 2
      IO_State_Cleaning : Byte;   // Status Reinigen
      IO_State_Testshot : Byte;   // Status Testschuss
      IO_Status : ANY;   // Status information of the robot interface
      IO_NewFault : Bool;
      IO_FaultLevel_1 : Bool;
      IO_FaultLevel_3 : Bool;
      IO_Faults : ANY;
   END_VAR
   VAR_TEMP
      Temp_IO_Status : "Fanuc_Status";   // Local status information of the robot interface
      Temp_IO_Fault : "Fanuc_Faults";   // Local fault information of the robot interface
      AnypointerStatus : ANY;   // Pointer for copying status information
      AnypointerFaults : ANY;   // Pointer for copying fault information
      LoopCounter : Int;   // Loopcounter
      NoOfMoulds : Byte;   // Number of moulds
      NoOfTimes : Byte;   // Number of times
      StartNecessary : Bool;   // Initial start of robot necessary
      PulsRobotInHomePos : Bool;   // Pulse robot in home position
      HFRobotInProgram : Bool;   // Help flag robot in program
      PulseNextShotTime : Bool;   // Puls for sending the next shot time to the robot
      TimeNo : Byte;   // Number of part shot in active mould
      RetValSFC : Int;
      TesShotSel_R1 : Bool;
      MaintProgSel_R1 : Bool;
      CleanProgSel_R1 : Bool;
   END_VAR
BEGIN

REGION Network 1: Load status information to local variables
         LAR1;
         L;
         LAR2;
   //
         L     W[AR2, P#0.0];  // Bytes
         T     W[AR1, P#0.0];
         L     W[AR2, P#2.0];  // Amount of bytes
         T     W[AR1, P#2.0];
         L     W[AR2, P#4.0];  // Block no,
         T     W[AR1, P#4.0];
         L     D[AR2, P#6.0];  // Startadress of data
         T     D[AR1, P#6.0];
         CALL  BLKMOV
         ( SRCBLK  := #AnypointerStatus,
           RET_VAL := #RetValSFC,
           DSTBLK  := #Temp_IO_Status
         );
   //
         LAR1;
         L;
         LAR2;
   //
         L     W[AR2, P#0.0];  // Bytes
         T     W[AR1, P#0.0];
         L     W[AR2, P#2.0];  // Amount of bytes
         T     W[AR1, P#2.0];
         L     W[AR2, P#4.0];  // Block no,
         T     W[AR1, P#4.0];
         L     D[AR2, P#6.0];  // Startadress of datas
         T     D[AR1, P#6.0];
         CALL  BLKMOV
         ( SRCBLK  := #AnypointerFaults,
           RET_VAL := #RetValSFC,
           DSTBLK  := #Temp_IO_Fault
         );

   // Read input data (outputs from robot)
         CALL  DPRD_DAT
         ( LADDR   := #IN_AdressRobIO,
           RET_VAL := #RetValSFC,
           RECORD  := #Temp_IO_Status.Output
         );
   //
END_REGION

REGION Network 2: Faults programm running from robot is missing
         A     #Temp_IO_Status.RequestAutomatic;
   //    UN    #Temp_Quit
         L     S5T#5S;
         SD    #IN_TimerDelayManSelect;  // #Timer_Prg_running
END_REGION

REGION Network 3: Fehler : Robot not for Datatransfer // FANUC
   //      UN    #Ext_Inputs_from_Robot.Ready_for_cycle
   //      U     #IN_Start_Prog_Imp
   //      ON    #Temp_IO_Status.Sys_Out.CMDENBL_Robot_ready
   //      O     #Temp_IO_Status.Sys_Out.Robot_Prg_paused
   //      U     #IN_Timer_Verz_Handanwahl   // #Timer_Prg_laeuft
   //      U     #IN_MK_Automatik
   //      =     #Status_Fanuc.Fault_Robot_not_ready
END_REGION

REGION Network 4: FAULT
         A     #IN_ResetFaultFct;
         R     #Temp_IO_Fault.FLT_System;
         R     #Temp_IO_Fault.FLT_Interface;
         R     #Temp_IO_Fault.FLT_Fuse_Supply;
   //
         A(;
         A     #IN_AutoStopOK;
         FP    #Temp_IO_Status.HfAutoStopOk;
         );
         A     #IN_MHAutomatic;
         A     #Temp_IO_Status.InterfaceOk;
         AN    #Temp_IO_Status.Input.diQuickStop;
         A     #Temp_IO_Status.InterfaceOk;
         O     #IN_ResetFaultFct;
         A     #Temp_IO_Status.Output.Fault_Robot;
         L     S5T#1S;
         SE    #IN_TimerFaultReset;
         A     #IN_TimerFaultReset;
         =     #Temp_IO_Status.Input.Robot_Fault_reset;
   //
   //      U     #IN_Reset_fault_Fkt
   //      U     #Temp_IO_Status.Output.doEmStop_Akt
   //      =     #Temp_IO_Status.Input.diResetEstop
   //
         A     #Temp_IO_Status.RequestAutomatic;
         A     #IN_TimerAutoOn;
         A     #Temp_IO_Status.Output.Fault_Robot;
         AN    #Temp_IO_Fault.FLT_System;
         S     #Temp_IO_Fault.FLT_System;
         S     #IO_NewFault;
         S     #IO_FaultLevel_1;
   //
         AN    #Temp_IO_Fault.FLT_System;
         AN    #Temp_IO_Fault.FLT_Interface;
         R     #Temp_IO_Status.FLT_detected;

         AN    #IN_FuseSupplyOK;
         S     #Temp_IO_Fault.FLT_Fuse_Supply;
   //
         O     #Temp_IO_Fault.FLT_System;
         O     #Temp_IO_Fault.FLT_Interface;
         A     #Temp_IO_Status.Output.CMDENBL_Robot_ready;
         A     #Temp_IO_Status.Output.SYSRDY_Robot_sys_ready;
         S     #Temp_IO_Status.FLT_detected;
   //
         AN    #Temp_IO_Status.FLT_detected;
         =     #Temp_IO_Status.InterfaceOk;

         L     #Temp_IO_Status.Output.GOError;
         T     #Temp_IO_Fault.FaultNumber;
END_REGION

REGION Network 5: Select auto/man requested
         A     #IN_ControlVoltage;
         A(;
         O     #IN_MHAutomatic;
         O     #Temp_IO_Status.Input.diHomeToMaintP;
         O     #Temp_IO_Status.Input.diMaintToHomeP;
         );
         A     #IN_AutoStopOK;
         AN    #IN_OtherRobotOnly;
   //    U     #Temp_IO_Status.Output.CMDENBL_Robot_ready
         A     #Temp_IO_Status.Output.SYSRDY_Robot_sys_ready;
         A     #Temp_IO_Status.InterfaceOk;
         AN(;
         A     #IN_ConfigWithTracking;
         A     #Temp_IO_Status.Output.doRobWaitWobj;
         AN    #IN_EnableFoamingCycle;
         A     #IN_TimerAutoOnTrack;
         );
         A     #Temp_IO_Status.Output.do_IRB_Auto;
         AN    #Temp_IO_Status.Input.diQuickStop;
         =     #Temp_IO_Status.RequestAutomatic;
   //
         AN    #Temp_IO_Status.RequestAutomatic;
         L     S5T#2S;
         SP    #IN_TimerAutoOFF;
   //
         A     #IN_TimerAutoOFF;
         CLR;
         ON    #IN_ControlVoltage;
         ON    #IN_AutoStopOK;
         ON    #IN_MHAutomatic;
         ON    #Temp_IO_Status.InterfaceOk;
         =     #Temp_IO_Status.RequestManualMode;
END_REGION

REGION Network 6: Decision how to start
         ON    #Temp_IO_Status.Output.CMDENBL_Robot_ready;
         ON    #Temp_IO_Status.Output.SYSRDY_Robot_sys_ready;
   //      O     #Temp_IO_Status.Output.doSysError
         S     #Temp_IO_Status.RobotNotInAuto;
   //
         O     #Temp_IO_Status.Output.doIRBInHome;
         FP    #Temp_IO_Status.FMRobotNotInAuto;
         =     #PulsRobotInHomePos;
         O     #Temp_IO_Status.Input.diStartCycle;
         O     #Temp_IO_Status.Input.diHomeToMaintP;
         O     #PulsRobotInHomePos;
         A     #Temp_IO_Status.Output.CMDENBL_Robot_ready;
         A     #Temp_IO_Status.Output.SYSRDY_Robot_sys_ready;
         R     #Temp_IO_Status.RobotNotInAuto;
   //
         A     #Temp_IO_Status.Output.doIRBInMaintP;
         O(;
         A     #Temp_IO_Status.Input.diBreak;
         AN    #Temp_IO_Status.Output.doIRBOutRangemc;
         );
         O(;
         A     #Temp_IO_Status.Input.diProgBreak;
         A     #Temp_IO_Status.Output.doIRBOutRangemc;
         );
         CLR;
         =     #HFRobotInProgram;
   //
         A     #HFRobotInProgram;
         AN    #Temp_IO_Status.RobotNotInAuto;
         AN(;
         A     #IN_ConfigWithTracking;
         A     #Temp_IO_Status.Output.doRobWaitWobj;
         );
         A     #Temp_IO_Status.RequestAutomatic;
         =     #Temp_IO_Status.RobotInProgram;
END_REGION

REGION Network 7: Roboter Positionen // MainPos, Reinigen
   // Während Zyklus Button ablöschen
         A     #IN_FoamingCycleRunning;
         AN    #Temp_IO_Status.Output.doIRBInHome;
         R     #IO_Button_MainPos;
         R     #IO_Button_Cleaning;

         A     #Temp_IO_Status.Output.Fault_Robot;
         R     #IO_Button_MainPos;

   // HomePos To MainPos
         A     #IO_Button_MainPos;
         AN    #IN_FoamingCycleRunning;
         A     #Temp_IO_Status.Output.doIRBInHome;
         A     #Temp_IO_Status.RequestAutomatic;
         JCN   MainPos;
         L     #IN_PGNO_MainPos;
         CAW;
         T     #Temp_IO_Status.Input.GIProgNo1;
         L     0;
         T     #Temp_IO_Status.Input.GIProgNo2;
         T     #Temp_IO_Status.Input.giTeachProgNo1;
         T     #Temp_IO_Status.Input.giTeachProgNo2;
         T     #Temp_IO_Status.Input.GIMCNo;

   MainPos:NOP   0;

   // HomePos to MainPos
         A     #IO_Button_MainPos;
         AN    #Temp_IO_Status.Output.doIRBInMaintP;
         A     #Temp_IO_Status.RequestAutomatic;
         =     #Temp_IO_Status.Input.diHomeToMaintP;